   RUNG wire#powerrail
      I_Contact( #Sensor_3 )
      I_Contact( "DB_Displacement".PlaceOcup.Sens3 )
   END_RUNG wire#w1
   RUNG wire#powerrail
      I_Contact( #Sensor_4 )
      I_Contact( "DB_Displacement".PlaceOcup.Sens4 )
   END_RUNG wire#w1
   // the same network as SCL:
   #Available := (NOT #Sensor_1 AND NOT "DB_Displacement".PlaceOcup.Sens1) OR (NOT #Sensor_2 AND NOT "DB_Displacement".PlaceOcup.Sens2) OR (NOT #Sensor_3 AND NOT "DB_Displacement".PlaceOcup.Sens3) OR (NOT #Sensor_4 AND NOT "DB_Displacement".PlaceOcup.Sens4);
END_REGION

REGION Network 2
   RUNG wire#powerrail
      Move(in := 280.0, out1 => #"Limit Y")
   END_RUNG
   // the same network as SCL:
   #"Limit Y" := 280.0;
END_REGION

REGION Network 3: Sensor 1 is not detect item
   RUNG wire#powerrail
      I_Contact( #Sensor_1 )
      I_Contact( "DB_Displacement".PlaceOcup.Sens1 )
      Move(in := 23.0, out1 => #"Ind Sensor_CO"."Sensor 1"."Pos X")
      Move(in := #"Limit Y", out1 => #"Ind Sensor_CO"."Sensor 1"."Pos Y")
      Move(in := 1, out1 => #"Ind Sensor_CO"."Sensor 1".SensorNumber)
      Move(in := #"Ind Sensor_CO"."Sensor 1", out1 => #"Sensor CO")
   END_RUNG
   // the same network as SCL:
   IF NOT #Sensor_1 AND NOT "DB_Displacement".PlaceOcup.Sens1 THEN
       #"Ind Sensor_CO"."Sensor 1"."Pos X" := 23.0;
       #"Ind Sensor_CO"."Sensor 1"."Pos Y" := #"Limit Y";
       #"Ind Sensor_CO"."Sensor 1".SensorNumber := 1;
       #"Sensor CO" := #"Ind Sensor_CO"."Sensor 1";
   END_IF;
END_REGION

REGION Network 4: Sensor 2 is not detect item
   RUNG wire#powerrail
      Contact( #Sensor_1 )
      wire#w1
      I_Contact( #Sensor_2 )
      I_Contact( "DB_Displacement".PlaceOcup.Sens2 )
      Move(in := 167.0, out1 => #"Ind Sensor_CO"."Sensor 2"."Pos X")
      Move(in := #"Limit Y", out1 => #"Ind Sensor_CO"."Sensor 2"."Pos Y")
      Move(in := 2, out1 => #"Ind Sensor_CO"."Sensor 2".SensorNumber)
      Move(in := #"Ind Sensor_CO"."Sensor 2", out1 => #"Sensor CO")
   END_RUNG
   RUNG wire#powerrail
      Contact( "DB_Displacement".PlaceOcup.Sens1 )
   END_RUNG wire#w1
   // the same network as SCL:
   IF (#Sensor_1 OR "DB_Displacement".PlaceOcup.Sens1) AND NOT #Sensor_2 AND NOT "DB_Displacement".PlaceOcup.Sens2 THEN
       #"Ind Sensor_CO"."Sensor 2"."Pos X" := 167.0;
       #"Ind Sensor_CO"."Sensor 2"."Pos Y" := #"Limit Y";
       #"Ind Sensor_CO"."Sensor 2".SensorNumber := 2;
       #"Sensor CO" := #"Ind Sensor_CO"."Sensor 2";
   END_IF;
END_REGION

REGION Network 5: Sensor 3 is not detect item
   RUNG wire#powerrail
      Contact( #Sensor_1 )
      wire#w1
      Contact( #Sensor_2 )
      wire#w2
      I_Contact( #Sensor_3 )
      wire#w3
      I_Contact( "DB_Displacement".PlaceOcup.Sens3 )
      Move(in := 313.0, out1 => #"Ind Sensor_CO"."Sensor 3"."Pos X")
      Move(in := #"Limit Y", out1 => #"Ind Sensor_CO"."Sensor 3"."Pos Y")
      Move(in := 3, out1 => #"Ind Sensor_CO"."Sensor 3".SensorNumber)
      Move(in := #"Ind Sensor_CO"."Sensor 3", out1 => #"Sensor CO")
   END_RUNG
   RUNG wire#powerrail
      Contact( "DB_Displacement".PlaceOcup.Sens1 )
   END_RUNG wire#w1
   RUNG wire#w1
      Contact( "DB_Displacement".PlaceOcup.Sens2 )
   END_RUNG wire#w2
   RUNG wire#w2
      Contact( "DB_Displacement".PlaceOcup.Sens3 )
   END_RUNG wire#w3
   // the same network as SCL:
   IF (#Sensor_1 OR "DB_Displacement".PlaceOcup.Sens1) AND (#Sensor_2 OR "DB_Displacement".PlaceOcup.Sens2) AND (NOT #Sensor_3 OR "DB_Displacement".PlaceOcup.Sens3) AND NOT "DB_Displacement".PlaceOcup.Sens3 THEN
       #"Ind Sensor_CO"."Sensor 3"."Pos X" := 313.0;
       #"Ind Sensor_CO"."Sensor 3"."Pos Y" := #"Limit Y";
       #"Ind Sensor_CO"."Sensor 3".SensorNumber := 3;
       #"Sensor CO" := #"Ind Sensor_CO"."Sensor 3";
   END_IF;
END_REGION

REGION Network 6: Sensor 4 is not detect item
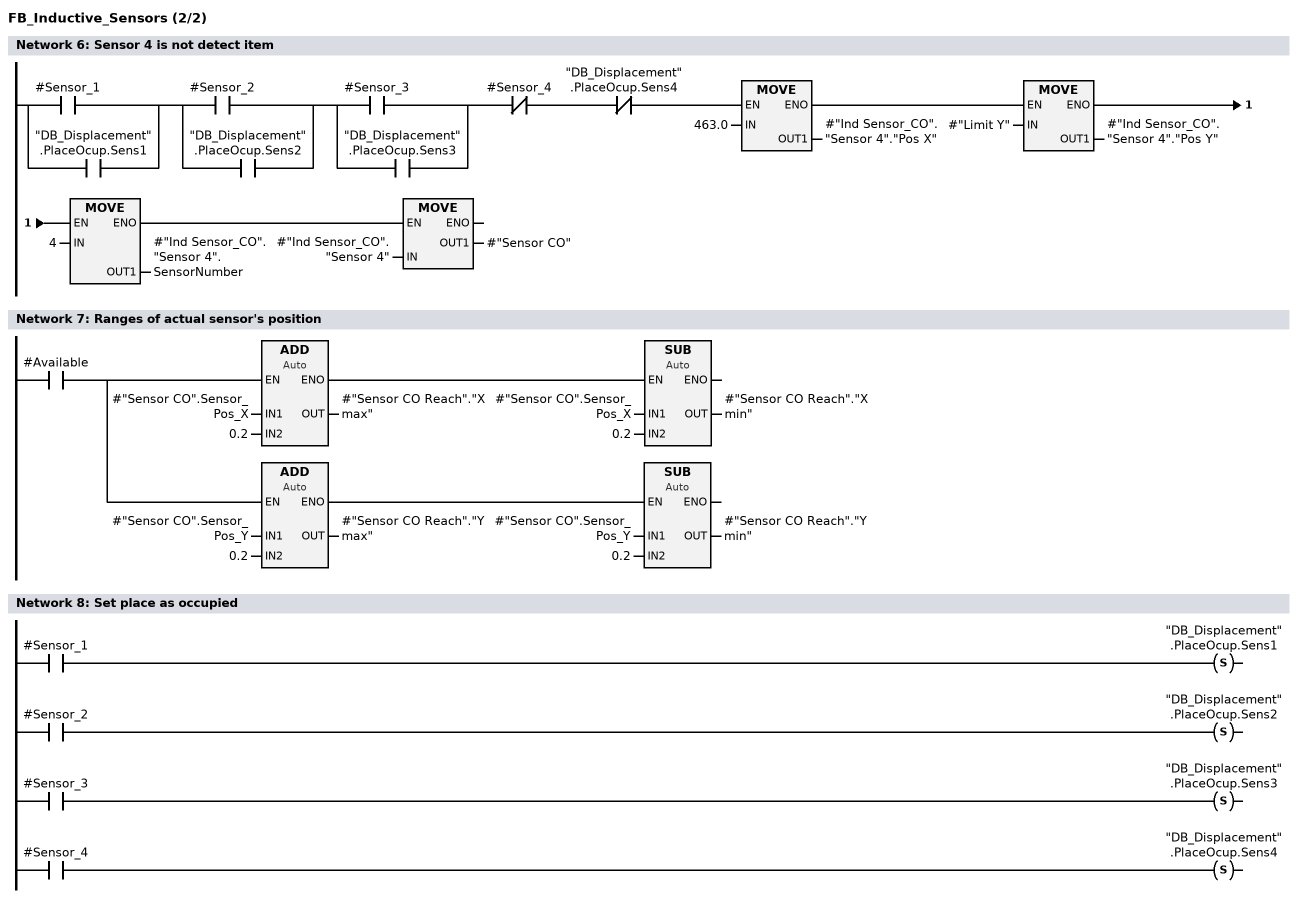
   RUNG wire#powerrail
      Contact( #Sensor_1 )
      wire#w1
      Contact( #Sensor_2 )
      wire#w2
      Contact( #Sensor_3 )
      wire#w3
      I_Contact( #Sensor_4 )
      I_Contact( "DB_Displacement".PlaceOcup.Sens4 )
      Move(in := 463.0, out1 => #"Ind Sensor_CO"."Sensor 4"."Pos X")
      Move(in := #"Limit Y", out1 => #"Ind Sensor_CO"."Sensor 4"."Pos Y")
      Move(in := 4, out1 => #"Ind Sensor_CO"."Sensor 4".SensorNumber)
      Move(in := #"Ind Sensor_CO"."Sensor 4", out1 => #"Sensor CO")
   END_RUNG
   RUNG wire#powerrail
      Contact( "DB_Displacement".PlaceOcup.Sens1 )
   END_RUNG wire#w1
   RUNG wire#w1
      Contact( "DB_Displacement".PlaceOcup.Sens2 )
   END_RUNG wire#w2
   RUNG wire#w2
      Contact( "DB_Displacement".PlaceOcup.Sens3 )
   END_RUNG wire#w3
   // the same network as SCL:
   IF (#Sensor_1 OR "DB_Displacement".PlaceOcup.Sens1) AND (#Sensor_2 OR "DB_Displacement".PlaceOcup.Sens2) AND (#Sensor_3 OR "DB_Displacement".PlaceOcup.Sens3) AND NOT #Sensor_4 AND NOT "DB_Displacement".PlaceOcup.Sens4 THEN
       #"Ind Sensor_CO"."Sensor 4"."Pos X" := 463.0;
       #"Ind Sensor_CO"."Sensor 4"."Pos Y" := #"Limit Y";
       #"Ind Sensor_CO"."Sensor 4".SensorNumber := 4;
       #"Sensor CO" := #"Ind Sensor_CO"."Sensor 4";
   END_IF;
END_REGION

REGION Network 7: Ranges of actual sensor's position
   RUNG wire#powerrail
      Contact( #Available )
      wire#w1
      Add(in1 := #"Sensor CO".Sensor_Pos_X, in2 := 0.2, out => #"Sensor CO Reach"."X max")
      Sub(in1 := #"Sensor CO".Sensor_Pos_X, in2 := 0.2, out => #"Sensor CO Reach"."X min")
   END_RUNG
   RUNG wire#w1
      Add(in1 := #"Sensor CO".Sensor_Pos_Y, in2 := 0.2, out => #"Sensor CO Reach"."Y max")
      Sub(in1 := #"Sensor CO".Sensor_Pos_Y, in2 := 0.2, out => #"Sensor CO Reach"."Y min")
   END_RUNG
   // the same network as SCL:
   IF #Available THEN
       #"Sensor CO Reach"."X max" := #"Sensor CO".Sensor_Pos_X + 0.2;
       #"Sensor CO Reach"."X min" := #"Sensor CO".Sensor_Pos_X - 0.2;
       #"Sensor CO Reach"."Y max" := #"Sensor CO".Sensor_Pos_Y + 0.2;
       #"Sensor CO Reach"."Y min" := #"Sensor CO".Sensor_Pos_Y - 0.2;
   END_IF;
END_REGION

REGION Network 8: Set place as occupied
   RUNG wire#powerrail
      Contact( #Sensor_1 )
      S_Coil( "DB_Displacement".PlaceOcup.Sens1 )
   END_RUNG
   RUNG wire#powerrail
      Contact( #Sensor_2 )
      S_Coil( "DB_Displacement".PlaceOcup.Sens2 )
   END_RUNG
   RUNG wire#powerrail
      Contact( #Sensor_3 )
      S_Coil( "DB_Displacement".PlaceOcup.Sens3 )
   END_RUNG
   RUNG wire#powerrail
      Contact( #Sensor_4 )
      S_Coil( "DB_Displacement".PlaceOcup.Sens4 )
   END_RUNG
   // the same network as SCL:
   IF #Sensor_1 THEN "DB_Displacement".PlaceOcup.Sens1 := TRUE; END_IF;
   IF #Sensor_2 THEN "DB_Displacement".PlaceOcup.Sens2 := TRUE; END_IF;
   IF #Sensor_3 THEN "DB_Displacement".PlaceOcup.Sens3 := TRUE; END_IF;
   IF #Sensor_4 THEN "DB_Displacement".PlaceOcup.Sens4 := TRUE; END_IF;
END_REGION
END_FUNCTION_BLOCK

// folder: Displacement/Object displacement/Velocity

FUNCTION_BLOCK "Velocity"   // FB16, LAD
{ S7_Optimized_Access := 'TRUE' }
VERSION : 0.1
   VAR_INPUT
      UDT_AxisStatus : Array[0..2] of "UDT_AxisStatus";
      TPx : Real;
      TPy : Real;
   END_VAR
   VAR_OUTPUT
      Vx : Real;
      Vy : Real;
   END_VAR
   VAR
      S : Real;
      HalfS : Real;
      Sx : Real;
      Sy : Real;
      Sx2 : Real;
      Sy2 : Real;
      Sum : Real;
      SPx : Real;
      SPy : Real;
      t : Real;
      SxActual : Real;
      Sx2Actual : Real;
      SyActual : Real;
      Sy2Actual : Real;
      SActual : Real;
      SumAct : Real;
      HalfSAct : Real;
   END_VAR
BEGIN

REGION Network 1
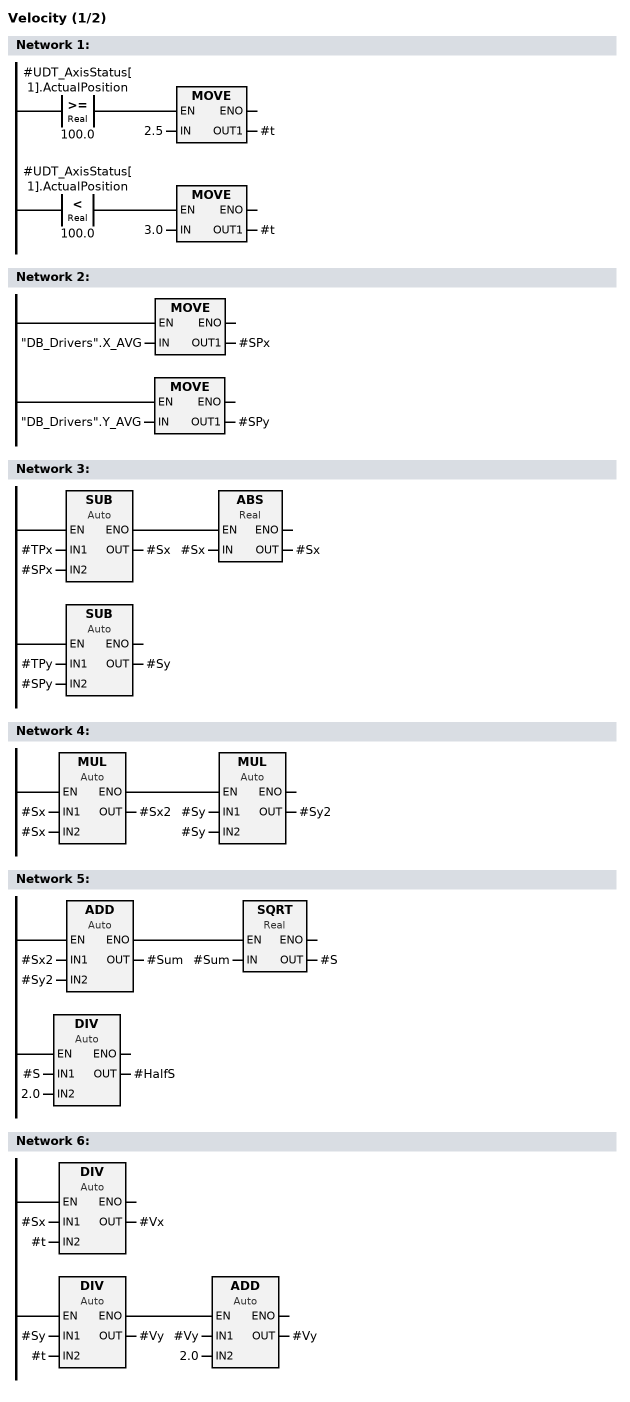
   RUNG wire#powerrail
      { S7_Templates := "SrcType := Real" } GE_Contact(in1 := #UDT_AxisStatus[1].ActualPosition, in2 := 100.0)
      Move(in := 2.5, out1 => #t)
   END_RUNG
   RUNG wire#powerrail
      { S7_Templates := "SrcType := Real" } LT_Contact(in1 := #UDT_AxisStatus[1].ActualPosition, in2 := 100.0)
      Move(in := 3.0, out1 => #t)
   END_RUNG
   // the same network as SCL:
   IF #UDT_AxisStatus[1].ActualPosition >= 100.0 THEN #t := 2.5; END_IF;
   IF #UDT_AxisStatus[1].ActualPosition < 100.0 THEN #t := 3.0; END_IF;
END_REGION

REGION Network 2
   RUNG wire#powerrail
      Move(in := "DB_Drivers".X_AVG, out1 => #SPx)
   END_RUNG
   RUNG wire#powerrail
      Move(in := "DB_Drivers".Y_AVG, out1 => #SPy)
   END_RUNG
   // the same network as SCL:
   #SPx := "DB_Drivers".X_AVG;
   #SPy := "DB_Drivers".Y_AVG;
END_REGION

REGION Network 3
   RUNG wire#powerrail
      Sub(in1 := #TPx, in2 := #SPx, out => #Sx)
      { S7_Templates := "SrcType := Real" } Abs(in := #Sx, out => #Sx)
   END_RUNG
   RUNG wire#powerrail
      Sub(in1 := #TPy, in2 := #SPy, out => #Sy)
   END_RUNG
   // the same network as SCL:
   #Sx := #TPx - #SPx;
   #Sx := ABS(#Sx);
   #Sy := #TPy - #SPy;
END_REGION

REGION Network 4
   RUNG wire#powerrail
      Mul(in1 := #Sx, in2 := #Sx, out => #Sx2)
      Mul(in1 := #Sy, in2 := #Sy, out => #Sy2)
   END_RUNG
   // the same network as SCL:
   #Sx2 := #Sx * #Sx;
   #Sy2 := #Sy * #Sy;
END_REGION

REGION Network 5
   #Sum := #Sx2 + #Sy2;
   #S := SQRT(#Sum);
   #HalfS := #S / 2.0;
END_REGION

REGION Network 6
   RUNG wire#powerrail
      Div(in1 := #Sx, in2 := #t, out => #Vx)
   END_RUNG
   RUNG wire#powerrail
      Div(in1 := #Sy, in2 := #t, out => #Vy)
      Add(in1 := #Vy, in2 := 2.0, out => #Vy)
   END_RUNG
   // the same network as SCL:
   #Vx := #Sx / #t;
   #Vy := #Sy / #t;
   #Vy := #Vy + 2.0;
END_REGION

REGION Network 7
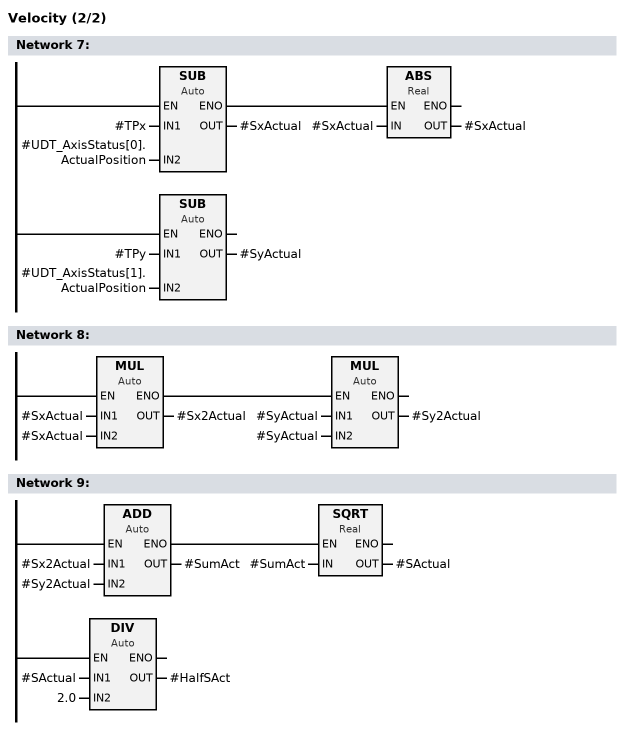
   RUNG wire#powerrail
      Sub(in1 := #TPx, in2 := #UDT_AxisStatus[0].ActualPosition, out => #SxActual)
      { S7_Templates := "SrcType := Real" } Abs(in := #SxActual, out => #SxActual)
   END_RUNG
   RUNG wire#powerrail
      Sub(in1 := #TPy, in2 := #UDT_AxisStatus[1].ActualPosition, out => #SyActual)
   END_RUNG
   // the same network as SCL:
   #SxActual := #TPx - #UDT_AxisStatus[0].ActualPosition;
   #SxActual := ABS(#SxActual);
   #SyActual := #TPy - #UDT_AxisStatus[1].ActualPosition;
END_REGION

REGION Network 8
   RUNG wire#powerrail
      Mul(in1 := #SxActual, in2 := #SxActual, out => #Sx2Actual)
      Mul(in1 := #SyActual, in2 := #SyActual, out => #Sy2Actual)
   END_RUNG
   // the same network as SCL:
   #Sx2Actual := #SxActual * #SxActual;
   #Sy2Actual := #SyActual * #SyActual;
END_REGION

REGION Network 9
   #SumAct := #Sx2Actual + #Sy2Actual;
   #SActual := SQRT(#SumAct);
   #HalfSAct := #SActual / 2.0;
END_REGION
END_FUNCTION_BLOCK

// folder: Drivers Parameters

FUNCTION_BLOCK "FB_Drivers"   // FB7, LAD
{ S7_Optimized_Access := 'TRUE' }
VERSION : 0.1
   VAR
      UDT_Axis_Control : Array[0..2] of "UDT_AxisControl";
      UDT_Axis_Status : Array[0..2] of "UDT_AxisStatus";
      X1 : Real;
      Y1 : Real;
      X2 : Real;
      Y2 : Real;
      X3 : Real;
      Y3 : Real;
      X4 : Real;
      Y4 : Real;
      X_AVG : Real;
      Y_AVG : Real;
   END_VAR
BEGIN

REGION Network 1: Axis Control
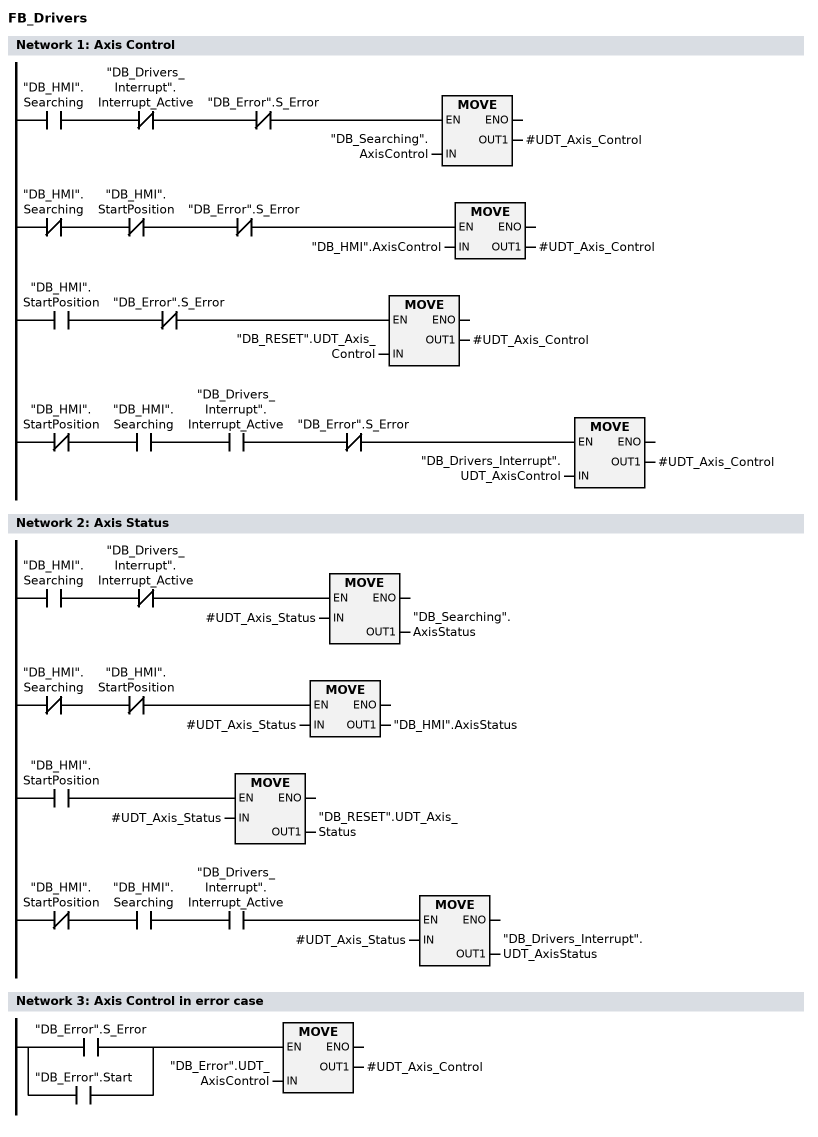
   RUNG wire#powerrail
      Contact( "DB_HMI".Searching )
      I_Contact( "DB_Drivers_Interrupt".Interrupt_Active )
      I_Contact( "DB_Error".S_Error )
      Move(in := "DB_Searching".AxisControl, out1 => #UDT_Axis_Control)
   END_RUNG
   RUNG wire#powerrail
      I_Contact( "DB_HMI".Searching )
      I_Contact( "DB_HMI".StartPosition )
      I_Contact( "DB_Error".S_Error )
      Move(in := "DB_HMI".AxisControl, out1 => #UDT_Axis_Control)
   END_RUNG
   RUNG wire#powerrail
      Contact( "DB_HMI".StartPosition )
      I_Contact( "DB_Error".S_Error )
      Move(in := "DB_RESET".UDT_Axis_Control, out1 => #UDT_Axis_Control)
   END_RUNG
   RUNG wire#powerrail
      I_Contact( "DB_HMI".StartPosition )
      Contact( "DB_HMI".Searching )
      Contact( "DB_Drivers_Interrupt".Interrupt_Active )
      I_Contact( "DB_Error".S_Error )
      Move(in := "DB_Drivers_Interrupt".UDT_AxisControl, out1 => #UDT_Axis_Control)
   END_RUNG
   // the same network as SCL:
   IF "DB_HMI".Searching AND NOT "DB_Drivers_Interrupt".Interrupt_Active AND NOT "DB_Error".S_Error THEN
       #UDT_Axis_Control := "DB_Searching".AxisControl;
   END_IF;
   IF NOT "DB_HMI".Searching AND NOT "DB_HMI".StartPosition AND NOT "DB_Error".S_Error THEN
       #UDT_Axis_Control := "DB_HMI".AxisControl;
   END_IF;
   IF "DB_HMI".StartPosition AND NOT "DB_Error".S_Error THEN
       #UDT_Axis_Control := "DB_RESET".UDT_Axis_Control;
   END_IF;
   IF NOT "DB_HMI".StartPosition AND "DB_HMI".Searching AND "DB_Drivers_Interrupt".Interrupt_Active AND NOT "DB_Error".S_Error THEN
       #UDT_Axis_Control := "DB_Drivers_Interrupt".UDT_AxisControl;
   END_IF;
END_REGION

REGION Network 2: Axis Status
   RUNG wire#powerrail
      Contact( "DB_HMI".Searching )
      I_Contact( "DB_Drivers_Interrupt".Interrupt_Active )
      Move(in := #UDT_Axis_Status, out1 => "DB_Searching".AxisStatus)
   END_RUNG
   RUNG wire#powerrail
      I_Contact( "DB_HMI".Searching )
      I_Contact( "DB_HMI".StartPosition )
      Move(in := #UDT_Axis_Status, out1 => "DB_HMI".AxisStatus)
   END_RUNG
   RUNG wire#powerrail
      Contact( "DB_HMI".StartPosition )
      Move(in := #UDT_Axis_Status, out1 => "DB_RESET".UDT_Axis_Status)
   END_RUNG
   RUNG wire#powerrail
      I_Contact( "DB_HMI".StartPosition )
      Contact( "DB_HMI".Searching )
      Contact( "DB_Drivers_Interrupt".Interrupt_Active )
      Move(in := #UDT_Axis_Status, out1 => "DB_Drivers_Interrupt".UDT_AxisStatus)
   END_RUNG
   // the same network as SCL:
   IF "DB_HMI".Searching AND NOT "DB_Drivers_Interrupt".Interrupt_Active THEN
       "DB_Searching".AxisStatus := #UDT_Axis_Status;
   END_IF;
   IF NOT "DB_HMI".Searching AND NOT "DB_HMI".StartPosition THEN
       "DB_HMI".AxisStatus := #UDT_Axis_Status;
   END_IF;
   IF "DB_HMI".StartPosition THEN "DB_RESET".UDT_Axis_Status := #UDT_Axis_Status; END_IF;
   IF NOT "DB_HMI".StartPosition AND "DB_HMI".Searching AND "DB_Drivers_Interrupt".Interrupt_Active THEN
       "DB_Drivers_Interrupt".UDT_AxisStatus := #UDT_Axis_Status;
   END_IF;
END_REGION

REGION Network 3: Axis Control in error case
   RUNG wire#powerrail
      Contact( "DB_Error".S_Error )
      wire#w1
      Move(in := "DB_Error".UDT_AxisControl, out1 => #UDT_Axis_Control)
   END_RUNG
   RUNG wire#powerrail
      Contact( "DB_Error".Start )
   END_RUNG wire#w1
   // the same network as SCL:
   IF "DB_Error".S_Error OR "DB_Error".Start THEN #UDT_Axis_Control := "DB_Error".UDT_AxisControl; END_IF;
END_REGION
END_FUNCTION_BLOCK

FUNCTION_BLOCK "FB_Drivers_Interrupt"   // FB12, LAD
{ S7_Optimized_Access := 'TRUE' }
VERSION : 0.1
   VAR
      Rising_IT_Counter : Int;   // Rising Edge Counter
      Falling_IT_Counter : Int;   // Falling Edge Counter
      UDT_AxisControl : Array[0..2] of "UDT_AxisControl";
      UDT_AxisStatus : Array[0..2] of "UDT_AxisStatus";   // Actual Axis Status
      Interrupt_Active : Bool;   // Item was detected. Interrupt is active.
      rtrig : Bool;   // rtrig connected with "stop" variable
      stop : Bool;   // Reset counters and variables when interrupt is done and target position is reached.
   END_VAR
   VAR CONSTANT
      false : Bool;
   END_VAR
BEGIN

REGION Network 1: Setting interrupt as active
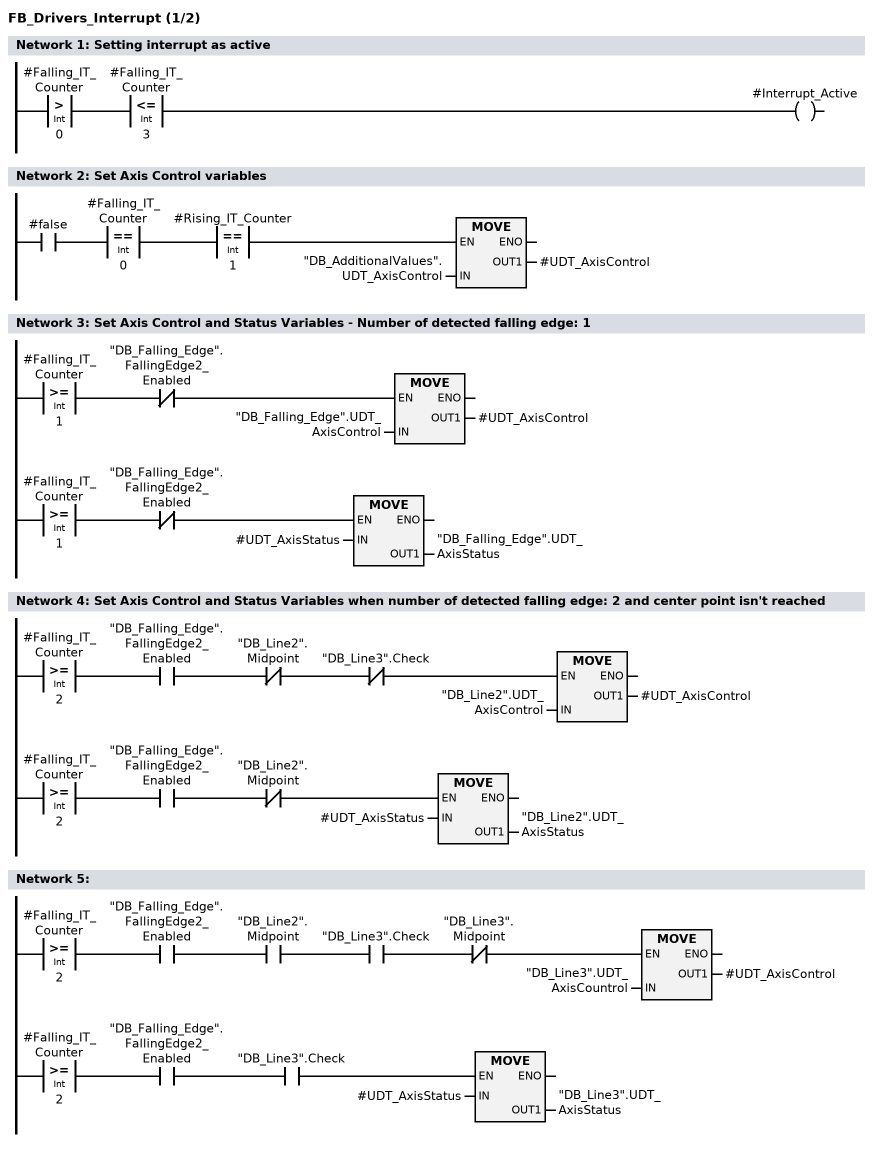
   RUNG wire#powerrail
      { S7_Templates := "SrcType := Int" } GT_Contact(in1 := #Falling_IT_Counter, in2 := 0)
      { S7_Templates := "SrcType := Int" } LE_Contact(in1 := #Falling_IT_Counter, in2 := 3)
      Coil( #Interrupt_Active )
   END_RUNG
   // the same network as SCL:
   #Interrupt_Active := (#Falling_IT_Counter > 0) AND (#Falling_IT_Counter <= 3);
END_REGION

REGION Network 2: Set Axis Control variables
   RUNG wire#powerrail
      Contact( #false )
      { S7_Templates := "SrcType := Int" } EQ_Contact(in1 := #Falling_IT_Counter, in2 := 0)
      { S7_Templates := "SrcType := Int" } EQ_Contact(in1 := #Rising_IT_Counter, in2 := 1)
      Move(in := "DB_AdditionalValues".UDT_AxisControl, out1 => #UDT_AxisControl)
   END_RUNG
   // the same network as SCL:
   IF #false AND (#Falling_IT_Counter = 0) AND (#Rising_IT_Counter = 1) THEN
       #UDT_AxisControl := "DB_AdditionalValues".UDT_AxisControl;
   END_IF;
END_REGION

REGION Network 3: Set Axis Control and Status Variables - Number of detected falling edge: 1
   RUNG wire#powerrail
      { S7_Templates := "SrcType := Int" } GE_Contact(in1 := #Falling_IT_Counter, in2 := 1)
      I_Contact( "DB_Falling_Edge".FallingEdge2_Enabled )
      Move(in := "DB_Falling_Edge".UDT_AxisControl, out1 => #UDT_AxisControl)
   END_RUNG
   RUNG wire#powerrail
      { S7_Templates := "SrcType := Int" } GE_Contact(in1 := #Falling_IT_Counter, in2 := 1)
      I_Contact( "DB_Falling_Edge".FallingEdge2_Enabled )
      Move(in := #UDT_AxisStatus, out1 => "DB_Falling_Edge".UDT_AxisStatus)
   END_RUNG
   // the same network as SCL:
   IF (#Falling_IT_Counter >= 1) AND NOT "DB_Falling_Edge".FallingEdge2_Enabled THEN
       #UDT_AxisControl := "DB_Falling_Edge".UDT_AxisControl;
       "DB_Falling_Edge".UDT_AxisStatus := #UDT_AxisStatus;
   END_IF;
END_REGION

REGION Network 4: Set Axis Control and Status Variables when number of detected falling edge: 2 and center point isn't reached
   RUNG wire#powerrail
      { S7_Templates := "SrcType := Int" } GE_Contact(in1 := #Falling_IT_Counter, in2 := 2)
      Contact( "DB_Falling_Edge".FallingEdge2_Enabled )
      I_Contact( "DB_Line2".Midpoint )
      I_Contact( "DB_Line3".Check )
      Move(in := "DB_Line2".UDT_AxisControl, out1 => #UDT_AxisControl)
   END_RUNG
   RUNG wire#powerrail
      { S7_Templates := "SrcType := Int" } GE_Contact(in1 := #Falling_IT_Counter, in2 := 2)
      Contact( "DB_Falling_Edge".FallingEdge2_Enabled )
      I_Contact( "DB_Line2".Midpoint )
      Move(in := #UDT_AxisStatus, out1 => "DB_Line2".UDT_AxisStatus)
   END_RUNG
   // the same network as SCL:
   IF (#Falling_IT_Counter >= 2) AND "DB_Falling_Edge".FallingEdge2_Enabled AND NOT "DB_Line2".Midpoint AND NOT "DB_Line3".Check THEN
       #UDT_AxisControl := "DB_Line2".UDT_AxisControl;
   END_IF;
   IF (#Falling_IT_Counter >= 2) AND "DB_Falling_Edge".FallingEdge2_Enabled AND NOT "DB_Line2".Midpoint THEN
       "DB_Line2".UDT_AxisStatus := #UDT_AxisStatus;
   END_IF;
END_REGION

REGION Network 5
   RUNG wire#powerrail
      { S7_Templates := "SrcType := Int" } GE_Contact(in1 := #Falling_IT_Counter, in2 := 2)
      Contact( "DB_Falling_Edge".FallingEdge2_Enabled )
      Contact( "DB_Line2".Midpoint )
      Contact( "DB_Line3".Check )
      I_Contact( "DB_Line3".Midpoint )
      Move(in := "DB_Line3".UDT_AxisCountrol, out1 => #UDT_AxisControl)
   END_RUNG
   RUNG wire#powerrail
      { S7_Templates := "SrcType := Int" } GE_Contact(in1 := #Falling_IT_Counter, in2 := 2)
      Contact( "DB_Falling_Edge".FallingEdge2_Enabled )
      Contact( "DB_Line3".Check )
      Move(in := #UDT_AxisStatus, out1 => "DB_Line3".UDT_AxisStatus)
   END_RUNG
   // the same network as SCL:
   IF (#Falling_IT_Counter >= 2) AND "DB_Falling_Edge".FallingEdge2_Enabled AND "DB_Line2".Midpoint AND "DB_Line3".Check AND NOT "DB_Line3".Midpoint THEN
       #UDT_AxisControl := "DB_Line3".UDT_AxisCountrol;
   END_IF;
   IF (#Falling_IT_Counter >= 2) AND "DB_Falling_Edge".FallingEdge2_Enabled AND "DB_Line3".Check THEN
       "DB_Line3".UDT_AxisStatus := #UDT_AxisStatus;
   END_IF;
END_REGION

REGION Network 6: Set Axis Control and Status Variables when center point is reached
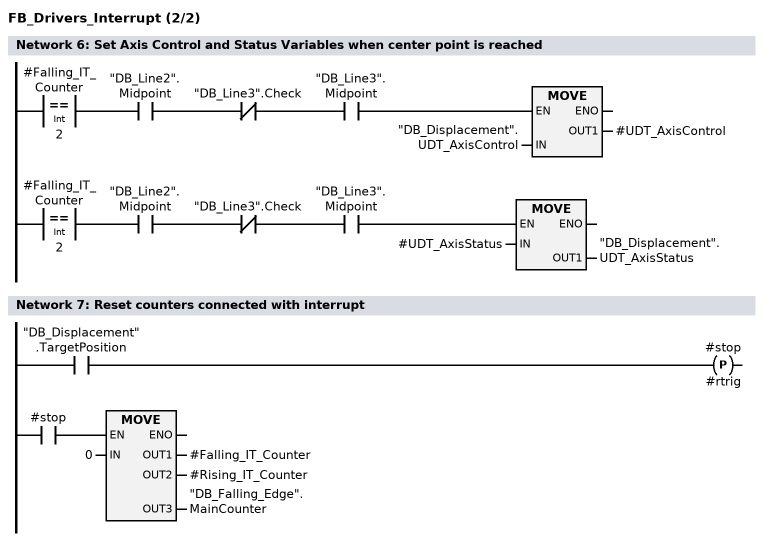
   RUNG wire#powerrail
      { S7_Templates := "SrcType := Int" } EQ_Contact(in1 := #Falling_IT_Counter, in2 := 2)
      Contact( "DB_Line2".Midpoint )
      I_Contact( "DB_Line3".Check )
      Contact( "DB_Line3".Midpoint )
      Move(in := "DB_Displacement".UDT_AxisControl, out1 => #UDT_AxisControl)
   END_RUNG
   RUNG wire#powerrail
      { S7_Templates := "SrcType := Int" } EQ_Contact(in1 := #Falling_IT_Counter, in2 := 2)
      Contact( "DB_Line2".Midpoint )
      I_Contact( "DB_Line3".Check )
      Contact( "DB_Line3".Midpoint )
      Move(in := #UDT_AxisStatus, out1 => "DB_Displacement".UDT_AxisStatus)
   END_RUNG
   // the same network as SCL:
   IF (#Falling_IT_Counter = 2) AND "DB_Line2".Midpoint AND NOT "DB_Line3".Check AND "DB_Line3".Midpoint THEN
       #UDT_AxisControl := "DB_Displacement".UDT_AxisControl;
       "DB_Displacement".UDT_AxisStatus := #UDT_AxisStatus;
   END_IF;
END_REGION

REGION Network 7: Reset counters connected with interrupt
   #stop := "DB_Displacement".TargetPosition AND NOT #rtrig;   // rising edge
   #rtrig := "DB_Displacement".TargetPosition;
   IF #stop THEN
       #Falling_IT_Counter := 0;
       #Rising_IT_Counter := 0;
       "DB_Falling_Edge".MainCounter := 0;
   END_IF;
END_REGION
END_FUNCTION_BLOCK

// folder: Electromagnet

FUNCTION "FC_Electromagnet" : Void   // FC1, LAD
{ S7_Optimized_Access := 'TRUE' }
VERSION : 0.1
BEGIN

REGION Network 1
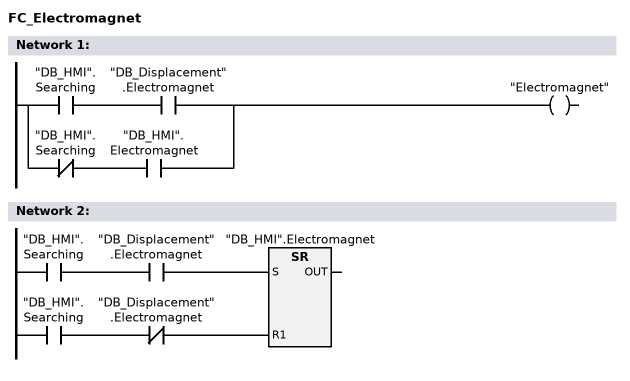
   RUNG wire#powerrail
      Contact( "DB_HMI".Searching )
      Contact( "DB_Displacement".Electromagnet )
      wire#w1
      Coil( "Electromagnet" )
   END_RUNG
   RUNG wire#powerrail
      I_Contact( "DB_HMI".Searching )
      Contact( "DB_HMI".Electromagnet )
   END_RUNG wire#w1
   // the same network as SCL:
   "Electromagnet" := ("DB_HMI".Searching AND "DB_Displacement".Electromagnet) OR (NOT "DB_HMI".Searching AND "DB_HMI".Electromagnet);
END_REGION

REGION Network 2
   RUNG wire#powerrail
      Contact( "DB_HMI".Searching )
      Contact( "DB_Displacement".Electromagnet )
      S_SR(operand := "DB_HMI".Electromagnet, r1 := wire#w1)
   END_RUNG
   RUNG wire#powerrail
      Contact( "DB_HMI".Searching )
      I_Contact( "DB_Displacement".Electromagnet )
   END_RUNG wire#w1
   // the same network as SCL:
   IF "DB_HMI".Searching AND "DB_Displacement".Electromagnet THEN
       "DB_HMI".Electromagnet := TRUE;   // SR flip-flop
   END_IF;
   IF "DB_HMI".Searching AND NOT "DB_Displacement".Electromagnet THEN
       "DB_HMI".Electromagnet := FALSE;
   END_IF;
END_REGION
END_FUNCTION

// folder: Error

FUNCTION_BLOCK "FB_Error"   // FB10, LAD
{ S7_Optimized_Access := 'TRUE' }
VERSION : 0.1
   VAR_INPUT
      Start : Bool;   // Reset error and start movement
   END_VAR
   VAR_OUTPUT
      "Error State" : Int;   // Set suitable color of error indicator
   END_VAR
   VAR_IN_OUT
      ResetError : Bool;   // Reset button
   END_VAR
   VAR
      Error : Bool;   // Active error
      UDT_AxisControl : Array[0..2] of "UDT_AxisControl";   // Axis Control variables
      UDT_AxisStatus : Array[0..2] of "UDT_AxisStatus";   // Axis Status variables
      S_Error : Bool;
      StartMoving : Bool;
      StartX : Bool;   // Start axis X movement
      PtrigX : Bool;   // Start axis X movement
      StartX2 : Bool;
      PtrigX2 : Bool;
      Ptrig : Bool;
      Set : Bool;
      PtrigReset : Bool;
      ResetValues : Bool;
      SetError : Bool;
      PtrigError : Bool;
      ItemToClose : Bool;
      DifY : Real;
      ErrorStateOne : Bool;
   END_VAR
   VAR_TEMP   // added for the SCL form of the ladder/FBD networks
      _w1 : Bool;
      _w2 : Bool;
   END_VAR
BEGIN

REGION Network 1